// TIA Portal project "CLU" (V13) (continued)
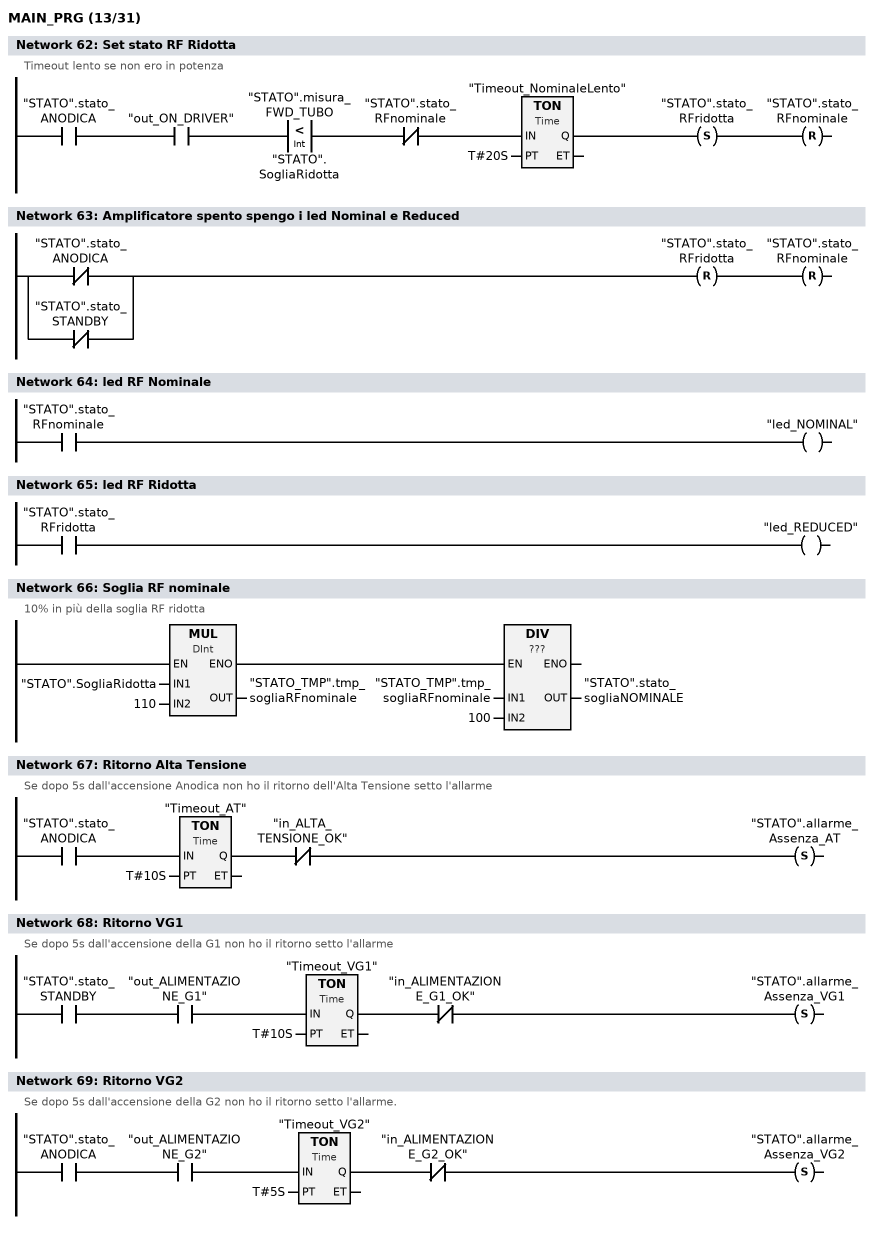
   "Timeout_NominaleLento".TON(IN := "STATO".stato_ANODICA AND "out_ON_DRIVER" AND ("STATO".misura_FWD_TUBO < "STATO".SogliaRidotta) AND NOT "STATO".stato_RFnominale,
                           PT := T#20S);
   IF "Timeout_NominaleLento".Q THEN
       "STATO".stato_RFridotta := TRUE;
       "STATO".stato_RFnominale := FALSE;
   END_IF;
END_REGION

REGION Network 63: Amplificatore spento spengo i led Nominal e Reduced
   RUNG wire#powerrail
      I_Contact( "STATO".stato_ANODICA )
      wire#w1
      R_Coil( "STATO".stato_RFridotta )
      R_Coil( "STATO".stato_RFnominale )
   END_RUNG
   RUNG wire#powerrail
      I_Contact( "STATO".stato_STANDBY )
   END_RUNG wire#w1
   // the same network as SCL:
   IF NOT "STATO".stato_ANODICA OR NOT "STATO".stato_STANDBY THEN
       "STATO".stato_RFridotta := FALSE;
       "STATO".stato_RFnominale := FALSE;
   END_IF;
END_REGION

REGION Network 64: led RF Nominale
   RUNG wire#powerrail
      Contact( "STATO".stato_RFnominale )
      Coil( "led_NOMINAL" )
   END_RUNG
   // the same network as SCL:
   "led_NOMINAL" := "STATO".stato_RFnominale;
END_REGION

REGION Network 65: led RF Ridotta
   RUNG wire#powerrail
      Contact( "STATO".stato_RFridotta )
      Coil( "led_REDUCED" )
   END_RUNG
   // the same network as SCL:
   "led_REDUCED" := "STATO".stato_RFridotta;
END_REGION

REGION Network 66: Soglia RF nominale
   // 10% in più della soglia RF ridotta
   RUNG wire#powerrail
      { S7_Templates := "SrcType := DInt" } Mul(in1 := "STATO".SogliaRidotta, in2 := 110, out => "STATO_TMP".tmp_sogliaRFnominale)
      { S7_Templates := "SrcType := ???" } Div(in1 := "STATO_TMP".tmp_sogliaRFnominale, in2 := 100, out => "STATO".stato_sogliaNOMINALE)
   END_RUNG
   // the same network as SCL:
   "STATO_TMP".tmp_sogliaRFnominale := "STATO".SogliaRidotta * 110;
   "STATO".stato_sogliaNOMINALE := "STATO_TMP".tmp_sogliaRFnominale / 100;
END_REGION

REGION Network 67: Ritorno Alta Tensione
   // Se dopo 5s dall'accensione Anodica non ho il ritorno dell'Alta Tensione setto l'allarme
   "Timeout_AT".TON(IN := "STATO".stato_ANODICA, PT := T#10S);
   IF "Timeout_AT".Q AND NOT "in_ALTA_TENSIONE_OK" THEN "STATO".allarme_Assenza_AT := TRUE; END_IF;
END_REGION

REGION Network 68: Ritorno VG1
   // Se dopo 5s dall'accensione della G1 non ho il ritorno setto l'allarme
   "Timeout_VG1".TON(IN := "STATO".stato_STANDBY AND "out_ALIMENTAZIONE_G1", PT := T#10S);
   IF "Timeout_VG1".Q AND NOT "in_ALIMENTAZIONE_G1_OK" THEN "STATO".allarme_Assenza_VG1 := TRUE; END_IF;
END_REGION

REGION Network 69: Ritorno VG2
   // Se dopo 5s dall'accensione della G2 non ho il ritorno setto l'allarme.
   "Timeout_VG2".TON(IN := "STATO".stato_ANODICA AND "out_ALIMENTAZIONE_G2", PT := T#5S);
   IF "Timeout_VG2".Q AND NOT "in_ALIMENTAZIONE_G2_OK" THEN "STATO".allarme_Assenza_VG2 := TRUE; END_IF;
END_REGION

REGION Network 70: Allarme mancanza VG1
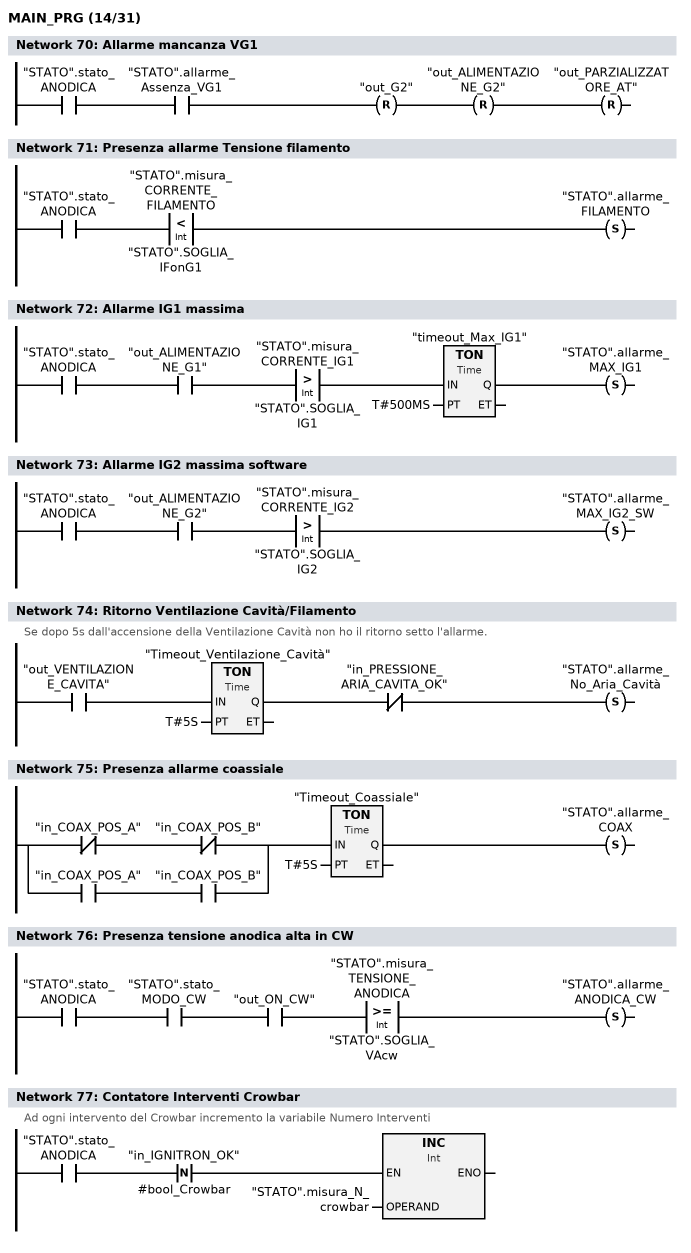
   RUNG wire#powerrail
      Contact( "STATO".stato_ANODICA )
      Contact( "STATO".allarme_Assenza_VG1 )
      R_Coil( "out_G2" )
      R_Coil( "out_ALIMENTAZIONE_G2" )
      R_Coil( "out_PARZIALIZZATORE_AT" )
   END_RUNG
   // the same network as SCL:
   IF "STATO".stato_ANODICA AND "STATO".allarme_Assenza_VG1 THEN
       "out_G2" := FALSE;
       "out_ALIMENTAZIONE_G2" := FALSE;
       "out_PARZIALIZZATORE_AT" := FALSE;
   END_IF;
END_REGION

REGION Network 71: Presenza allarme Tensione filamento
   RUNG wire#powerrail
      Contact( "STATO".stato_ANODICA )
      { S7_Templates := "SrcType := Int" } LT_Contact(in1 := "STATO".misura_CORRENTE_FILAMENTO, in2 := "STATO".SOGLIA_IFonG1)
      S_Coil( "STATO".allarme_FILAMENTO )
   END_RUNG
   // the same network as SCL:
   IF "STATO".stato_ANODICA AND ("STATO".misura_CORRENTE_FILAMENTO < "STATO".SOGLIA_IFonG1) THEN
       "STATO".allarme_FILAMENTO := TRUE;
   END_IF;
END_REGION

REGION Network 72: Allarme IG1 massima
   "timeout_Max_IG1".TON(IN := "STATO".stato_ANODICA AND "out_ALIMENTAZIONE_G1" AND ("STATO".misura_CORRENTE_IG1 > "STATO".SOGLIA_IG1),
                         PT := T#500MS);
   IF "timeout_Max_IG1".Q THEN "STATO".allarme_MAX_IG1 := TRUE; END_IF;
END_REGION

REGION Network 73: Allarme IG2 massima software
   RUNG wire#powerrail
      Contact( "STATO".stato_ANODICA )
      Contact( "out_ALIMENTAZIONE_G2" )
      { S7_Templates := "SrcType := Int" } GT_Contact(in1 := "STATO".misura_CORRENTE_IG2, in2 := "STATO".SOGLIA_IG2)
      S_Coil( "STATO".allarme_MAX_IG2_SW )
   END_RUNG
   // the same network as SCL:
   IF "STATO".stato_ANODICA AND "out_ALIMENTAZIONE_G2" AND ("STATO".misura_CORRENTE_IG2 > "STATO".SOGLIA_IG2) THEN
       "STATO".allarme_MAX_IG2_SW := TRUE;
   END_IF;
END_REGION

REGION Network 74: Ritorno Ventilazione Cavità/Filamento
   // Se dopo 5s dall'accensione della Ventilazione Cavità non ho il ritorno setto l'allarme.
   "Timeout_Ventilazione_Cavità".TON(IN := "out_VENTILAZIONE_CAVITA", PT := T#5S);
   IF "Timeout_Ventilazione_Cavità".Q AND NOT "in_PRESSIONE_ARIA_CAVITA_OK" THEN
       "STATO".allarme_No_Aria_Cavità := TRUE;
   END_IF;
END_REGION

REGION Network 75: Presenza allarme coassiale
   "Timeout_Coassiale".TON(IN := (NOT "in_COAX_POS_A" AND NOT "in_COAX_POS_B") OR ("in_COAX_POS_A" AND "in_COAX_POS_B"),
                           PT := T#5S);
   IF "Timeout_Coassiale".Q THEN "STATO".allarme_COAX := TRUE; END_IF;
END_REGION

REGION Network 76: Presenza tensione anodica alta in CW
   RUNG wire#powerrail
      Contact( "STATO".stato_ANODICA )
      Contact( "STATO".stato_MODO_CW )
      Contact( "out_ON_CW" )
      { S7_Templates := "SrcType := Int" } GE_Contact(in1 := "STATO".misura_TENSIONE_ANODICA, in2 := "STATO".SOGLIA_VAcw)
      S_Coil( "STATO".allarme_ANODICA_CW )
   END_RUNG
   // the same network as SCL:
   IF "STATO".stato_ANODICA AND "STATO".stato_MODO_CW AND "out_ON_CW" AND ("STATO".misura_TENSIONE_ANODICA >= "STATO".SOGLIA_VAcw) THEN
       "STATO".allarme_ANODICA_CW := TRUE;
   END_IF;
END_REGION

REGION Network 77: Contatore Interventi Crowbar
   // Ad ogni intervento del Crowbar incremento la variabile Numero Interventi
   RUNG wire#powerrail
      Contact( "STATO".stato_ANODICA )
      N_Contact(operand := "in_IGNITRON_OK", bit := #bool_Crowbar)
      { S7_Templates := "DestType := Int" } Inc( "STATO".misura_N_crowbar )
   END_RUNG
   // the same network as SCL:
   #_w1 := "STATO".stato_ANODICA AND NOT "in_IGNITRON_OK" AND #bool_Crowbar;   // falling edge of "in_IGNITRON_OK"
   #bool_Crowbar := "in_IGNITRON_OK";
   IF #_w1 THEN "STATO".misura_N_crowbar := "STATO".misura_N_crowbar + 1; END_IF;
END_REGION

REGION Network 78: Soglia ROS 400kW
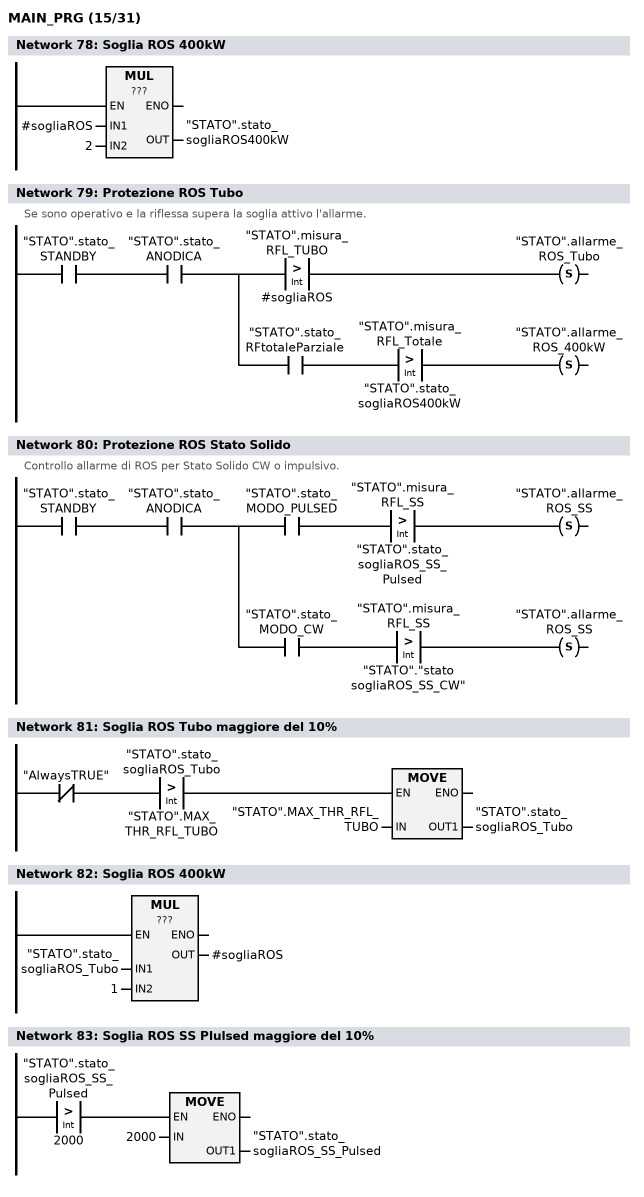
   RUNG wire#powerrail
      { S7_Templates := "SrcType := ???" } Mul(in1 := #sogliaROS, in2 := 2, out => "STATO".stato_sogliaROS400kW)
   END_RUNG
   // the same network as SCL:
   "STATO".stato_sogliaROS400kW := #sogliaROS * 2;
END_REGION

REGION Network 79: Protezione ROS Tubo
   // Se sono operativo e la riflessa supera la soglia attivo l'allarme.
   RUNG wire#powerrail
      Contact( "STATO".stato_STANDBY )
      Contact( "STATO".stato_ANODICA )
      wire#w1
      { S7_Templates := "SrcType := Int" } GT_Contact(in1 := "STATO".misura_RFL_TUBO, in2 := #sogliaROS)
      S_Coil( "STATO".allarme_ROS_Tubo )
   END_RUNG
   RUNG wire#w1
      Contact( "STATO".stato_RFtotaleParziale )
      { S7_Templates := "SrcType := Int" } GT_Contact(in1 := "STATO".misura_RFL_Totale, in2 := "STATO".stato_sogliaROS400kW)
      S_Coil( "STATO".allarme_ROS_400kW )
   END_RUNG
   // the same network as SCL:
   #_w1 := "STATO".stato_STANDBY AND "STATO".stato_ANODICA;
   IF #_w1 AND ("STATO".misura_RFL_TUBO > #sogliaROS) THEN "STATO".allarme_ROS_Tubo := TRUE; END_IF;
   IF #_w1 AND "STATO".stato_RFtotaleParziale AND ("STATO".misura_RFL_Totale > "STATO".stato_sogliaROS400kW) THEN
       "STATO".allarme_ROS_400kW := TRUE;
   END_IF;
END_REGION

REGION Network 80: Protezione ROS Stato Solido
   // Controllo allarme di ROS per Stato Solido CW o impulsivo.
   RUNG wire#powerrail
      Contact( "STATO".stato_STANDBY )
      Contact( "STATO".stato_ANODICA )
      wire#w1
      Contact( "STATO".stato_MODO_PULSED )
      { S7_Templates := "SrcType := Int" } GT_Contact(in1 := "STATO".misura_RFL_SS, in2 := "STATO".stato_sogliaROS_SS_Pulsed)
      S_Coil( "STATO".allarme_ROS_SS )
   END_RUNG
   RUNG wire#w1
      Contact( "STATO".stato_MODO_CW )
      { S7_Templates := "SrcType := Int" } GT_Contact(in1 := "STATO".misura_RFL_SS, in2 := "STATO"."stato sogliaROS_SS_CW")
      S_Coil( "STATO".allarme_ROS_SS )
   END_RUNG
   // the same network as SCL:
   #_w1 := "STATO".stato_STANDBY AND "STATO".stato_ANODICA;
   IF #_w1 AND "STATO".stato_MODO_PULSED AND ("STATO".misura_RFL_SS > "STATO".stato_sogliaROS_SS_Pulsed) THEN
       "STATO".allarme_ROS_SS := TRUE;
   END_IF;
   IF #_w1 AND "STATO".stato_MODO_CW AND ("STATO".misura_RFL_SS > "STATO"."stato sogliaROS_SS_CW") THEN
       "STATO".allarme_ROS_SS := TRUE;
   END_IF;
END_REGION

REGION Network 81: Soglia ROS Tubo maggiore del 10%
   RUNG wire#powerrail
      I_Contact( "AlwaysTRUE" )
      { S7_Templates := "SrcType := Int" } GT_Contact(in1 := "STATO".stato_sogliaROS_Tubo, in2 := "STATO".MAX_THR_RFL_TUBO)
      Move(in := "STATO".MAX_THR_RFL_TUBO, out1 => "STATO".stato_sogliaROS_Tubo)
   END_RUNG
   // the same network as SCL:
   IF NOT "AlwaysTRUE" AND ("STATO".stato_sogliaROS_Tubo > "STATO".MAX_THR_RFL_TUBO) THEN
       "STATO".stato_sogliaROS_Tubo := "STATO".MAX_THR_RFL_TUBO;
   END_IF;
END_REGION

REGION Network 82: Soglia ROS 400kW
   RUNG wire#powerrail
      { S7_Templates := "SrcType := ???" } Mul(in1 := "STATO".stato_sogliaROS_Tubo, in2 := 1, out => #sogliaROS)
   END_RUNG
   // the same network as SCL:
   #sogliaROS := "STATO".stato_sogliaROS_Tubo * 1;
END_REGION

REGION Network 83: Soglia ROS SS Plulsed maggiore del 10%
   RUNG wire#powerrail
      { S7_Templates := "SrcType := Int" } GT_Contact(in1 := "STATO".stato_sogliaROS_SS_Pulsed, in2 := 2000)
      Move(in := 2000, out1 => "STATO".stato_sogliaROS_SS_Pulsed)
   END_RUNG
   // the same network as SCL:
   IF "STATO".stato_sogliaROS_SS_Pulsed > 2000 THEN "STATO".stato_sogliaROS_SS_Pulsed := 2000; END_IF;
END_REGION

REGION Network 84: Soglia ROS SS CW maggiore del 10%
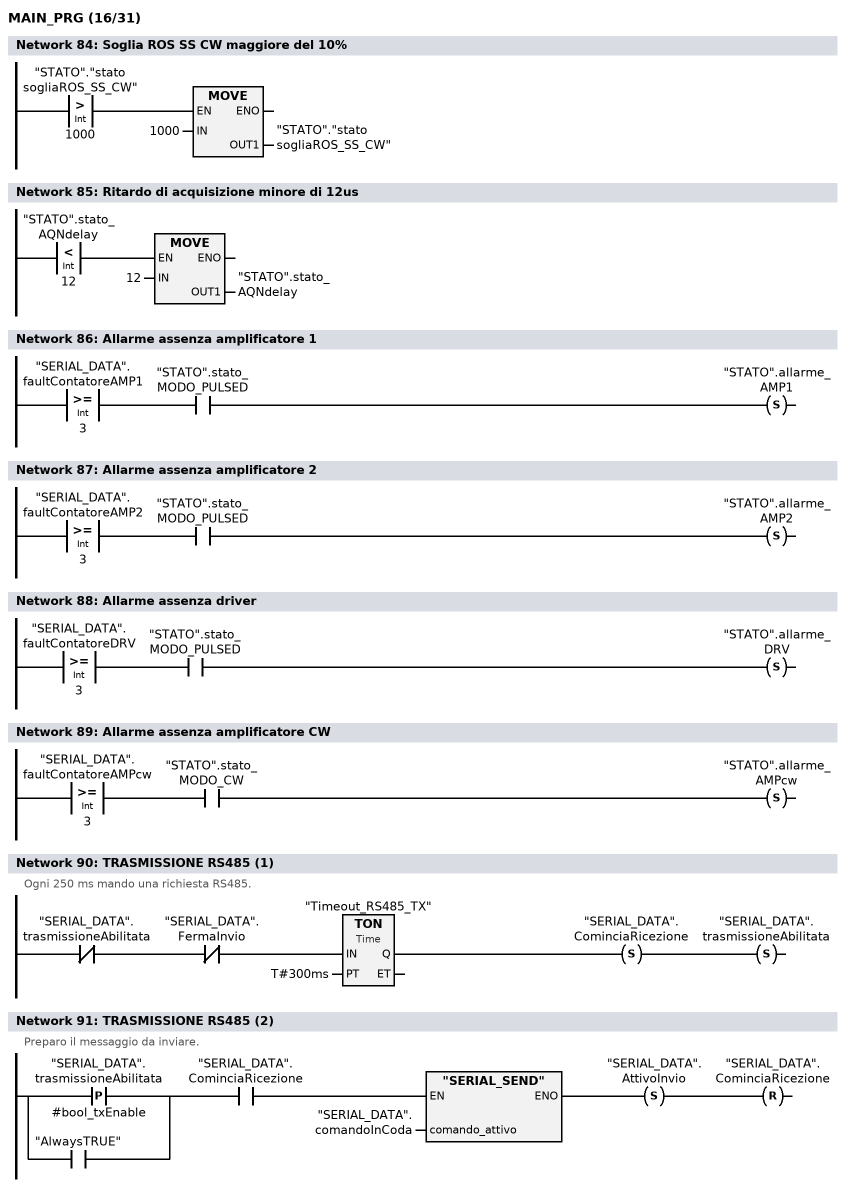
   RUNG wire#powerrail
      { S7_Templates := "SrcType := Int" } GT_Contact(in1 := "STATO"."stato sogliaROS_SS_CW", in2 := 1000)
      Move(in := 1000, out1 => "STATO"."stato sogliaROS_SS_CW")
   END_RUNG
   // the same network as SCL:
   IF "STATO"."stato sogliaROS_SS_CW" > 1000 THEN "STATO"."stato sogliaROS_SS_CW" := 1000; END_IF;
END_REGION

REGION Network 85: Ritardo di acquisizione minore di 12us
   RUNG wire#powerrail
      { S7_Templates := "SrcType := Int" } LT_Contact(in1 := "STATO".stato_AQNdelay, in2 := 12)
      Move(in := 12, out1 => "STATO".stato_AQNdelay)
   END_RUNG
   // the same network as SCL:
   IF "STATO".stato_AQNdelay < 12 THEN "STATO".stato_AQNdelay := 12; END_IF;
END_REGION

REGION Network 86: Allarme assenza amplificatore 1
   RUNG wire#powerrail
      { S7_Templates := "SrcType := Int" } GE_Contact(in1 := "SERIAL_DATA".faultContatoreAMP1, in2 := 3)
      Contact( "STATO".stato_MODO_PULSED )
      S_Coil( "STATO".allarme_AMP1 )
   END_RUNG
   // the same network as SCL:
   IF ("SERIAL_DATA".faultContatoreAMP1 >= 3) AND "STATO".stato_MODO_PULSED THEN
       "STATO".allarme_AMP1 := TRUE;
   END_IF;
END_REGION

REGION Network 87: Allarme assenza amplificatore 2
   RUNG wire#powerrail
      { S7_Templates := "SrcType := Int" } GE_Contact(in1 := "SERIAL_DATA".faultContatoreAMP2, in2 := 3)
      Contact( "STATO".stato_MODO_PULSED )
      S_Coil( "STATO".allarme_AMP2 )
   END_RUNG
   // the same network as SCL:
   IF ("SERIAL_DATA".faultContatoreAMP2 >= 3) AND "STATO".stato_MODO_PULSED THEN
       "STATO".allarme_AMP2 := TRUE;
   END_IF;
END_REGION

REGION Network 88: Allarme assenza driver
   RUNG wire#powerrail
      { S7_Templates := "SrcType := Int" } GE_Contact(in1 := "SERIAL_DATA".faultContatoreDRV, in2 := 3)
      Contact( "STATO".stato_MODO_PULSED )
      S_Coil( "STATO".allarme_DRV )
   END_RUNG
   // the same network as SCL:
   IF ("SERIAL_DATA".faultContatoreDRV >= 3) AND "STATO".stato_MODO_PULSED THEN
       "STATO".allarme_DRV := TRUE;
   END_IF;
END_REGION

REGION Network 89: Allarme assenza amplificatore CW
   RUNG wire#powerrail
      { S7_Templates := "SrcType := Int" } GE_Contact(in1 := "SERIAL_DATA".faultContatoreAMPcw, in2 := 3)
      Contact( "STATO".stato_MODO_CW )
      S_Coil( "STATO".allarme_AMPcw )
   END_RUNG
   // the same network as SCL:
   IF ("SERIAL_DATA".faultContatoreAMPcw >= 3) AND "STATO".stato_MODO_CW THEN
       "STATO".allarme_AMPcw := TRUE;
   END_IF;
END_REGION

REGION Network 90: TRASMISSIONE RS485 (1)
   // Ogni 250 ms mando una richiesta RS485.
   "Timeout_RS485_TX".TON(IN := NOT "SERIAL_DATA".trasmissioneAbilitata AND NOT "SERIAL_DATA".FermaInvio,
                          PT := T#300ms);
   IF "Timeout_RS485_TX".Q THEN
       "SERIAL_DATA".CominciaRicezione := TRUE;
       "SERIAL_DATA".trasmissioneAbilitata := TRUE;
   END_IF;
END_REGION

REGION Network 91: TRASMISSIONE RS485 (2)
   // Preparo il messaggio da inviare.
   RUNG wire#powerrail
      P_Contact(operand := "SERIAL_DATA".trasmissioneAbilitata, bit := #bool_txEnable)
      wire#w1
      Contact( "SERIAL_DATA".CominciaRicezione )
      "SERIAL_SEND"(comando_attivo := "SERIAL_DATA".comandoInCoda)
      S_Coil( "SERIAL_DATA".AttivoInvio )
      R_Coil( "SERIAL_DATA".CominciaRicezione )
   END_RUNG
   RUNG wire#powerrail
      Contact( "AlwaysTRUE" )
   END_RUNG wire#w1
   // the same network as SCL:
   #_w1 := "SERIAL_DATA".trasmissioneAbilitata AND NOT #bool_txEnable;   // rising edge of "SERIAL_DATA".trasmissioneAbilitata
   #bool_txEnable := "SERIAL_DATA".trasmissioneAbilitata;
   "SERIAL_SEND"(EN := (#_w1 OR "AlwaysTRUE") AND "SERIAL_DATA".CominciaRicezione,
                 comando_attivo := "SERIAL_DATA".comandoInCoda,
                 ENO => #_w2);
   IF #_w2 THEN
       "SERIAL_DATA".AttivoInvio := TRUE;
       "SERIAL_DATA".CominciaRicezione := FALSE;
   END_IF;
END_REGION

REGION Network 92: TRASMISSIONE RS485 (3): 76h
   // Processo la richiesta di stato ID==0
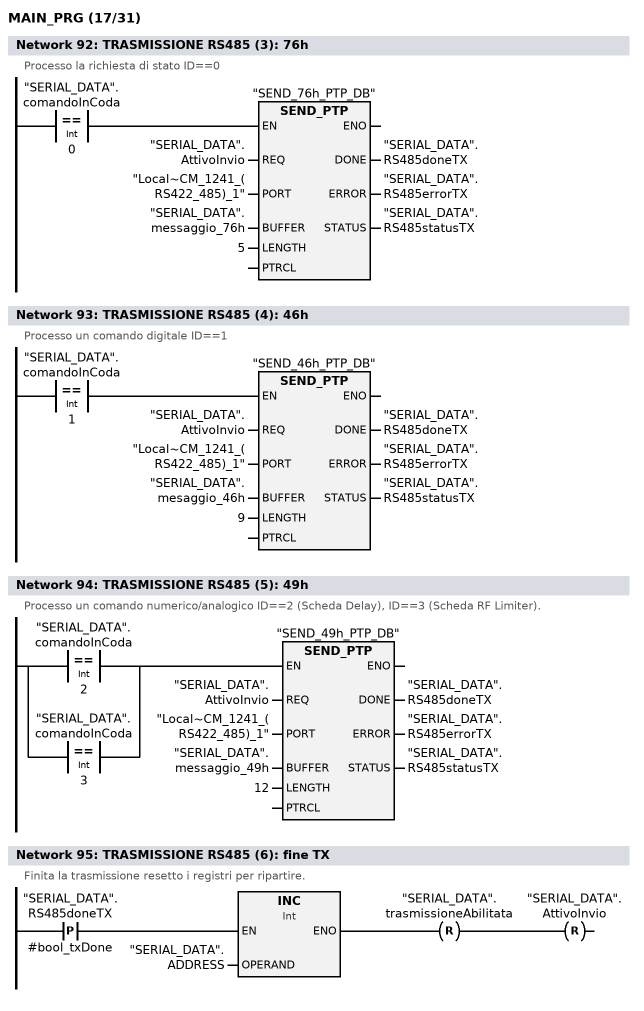
   IF "SERIAL_DATA".comandoInCoda = 0 THEN
       "SEND_76h_PTP_DB"(REQ := "SERIAL_DATA".AttivoInvio,   // SEND_PTP
                         PORT := "Local~CM_1241_(RS422_485)_1",
                         BUFFER := "SERIAL_DATA".messaggio_76h,
                         LENGTH := 5,
                         DONE => "SERIAL_DATA".RS485doneTX,
                         ERROR => "SERIAL_DATA".RS485errorTX,
                         STATUS => "SERIAL_DATA".RS485statusTX);
   END_IF;
END_REGION

REGION Network 93: TRASMISSIONE RS485 (4): 46h
   // Processo un comando digitale ID==1
   IF "SERIAL_DATA".comandoInCoda = 1 THEN
       "SEND_46h_PTP_DB"(REQ := "SERIAL_DATA".AttivoInvio,   // SEND_PTP
                         PORT := "Local~CM_1241_(RS422_485)_1",
                         BUFFER := "SERIAL_DATA".mesaggio_46h,
                         LENGTH := 9,
                         DONE => "SERIAL_DATA".RS485doneTX,
                         ERROR => "SERIAL_DATA".RS485errorTX,
                         STATUS => "SERIAL_DATA".RS485statusTX);
   END_IF;
END_REGION

REGION Network 94: TRASMISSIONE RS485 (5): 49h
   // Processo un comando numerico/analogico ID==2 (Scheda Delay), ID==3 (Scheda RF Limiter).
   IF ("SERIAL_DATA".comandoInCoda = 2) OR ("SERIAL_DATA".comandoInCoda = 3) THEN
       "SEND_49h_PTP_DB"(REQ := "SERIAL_DATA".AttivoInvio,   // SEND_PTP
                         PORT := "Local~CM_1241_(RS422_485)_1",
                         BUFFER := "SERIAL_DATA".messaggio_49h,
                         LENGTH := 12,
                         DONE => "SERIAL_DATA".RS485doneTX,
                         ERROR => "SERIAL_DATA".RS485errorTX,
                         STATUS => "SERIAL_DATA".RS485statusTX);
   END_IF;
END_REGION

REGION Network 95: TRASMISSIONE RS485 (6): fine TX
   // Finita la trasmissione resetto i registri per ripartire.
   RUNG wire#powerrail
      P_Contact(operand := "SERIAL_DATA".RS485doneTX, bit := #bool_txDone)
      { S7_Templates := "DestType := Int" } Inc( "SERIAL_DATA".ADDRESS )
      R_Coil( "SERIAL_DATA".trasmissioneAbilitata )
      R_Coil( "SERIAL_DATA".AttivoInvio )
   END_RUNG
   // the same network as SCL:
   #_w1 := "SERIAL_DATA".RS485doneTX AND NOT #bool_txDone;   // rising edge of "SERIAL_DATA".RS485doneTX
   #bool_txDone := "SERIAL_DATA".RS485doneTX;
   IF #_w1 THEN
       "SERIAL_DATA".ADDRESS := "SERIAL_DATA".ADDRESS + 1;
       "SERIAL_DATA".trasmissioneAbilitata := FALSE;
       "SERIAL_DATA".AttivoInvio := FALSE;
   END_IF;
END_REGION

REGION Network 96: RICEZIONE RS485 (1): ricezione
   // La ricezione seriale è sempre attiva.
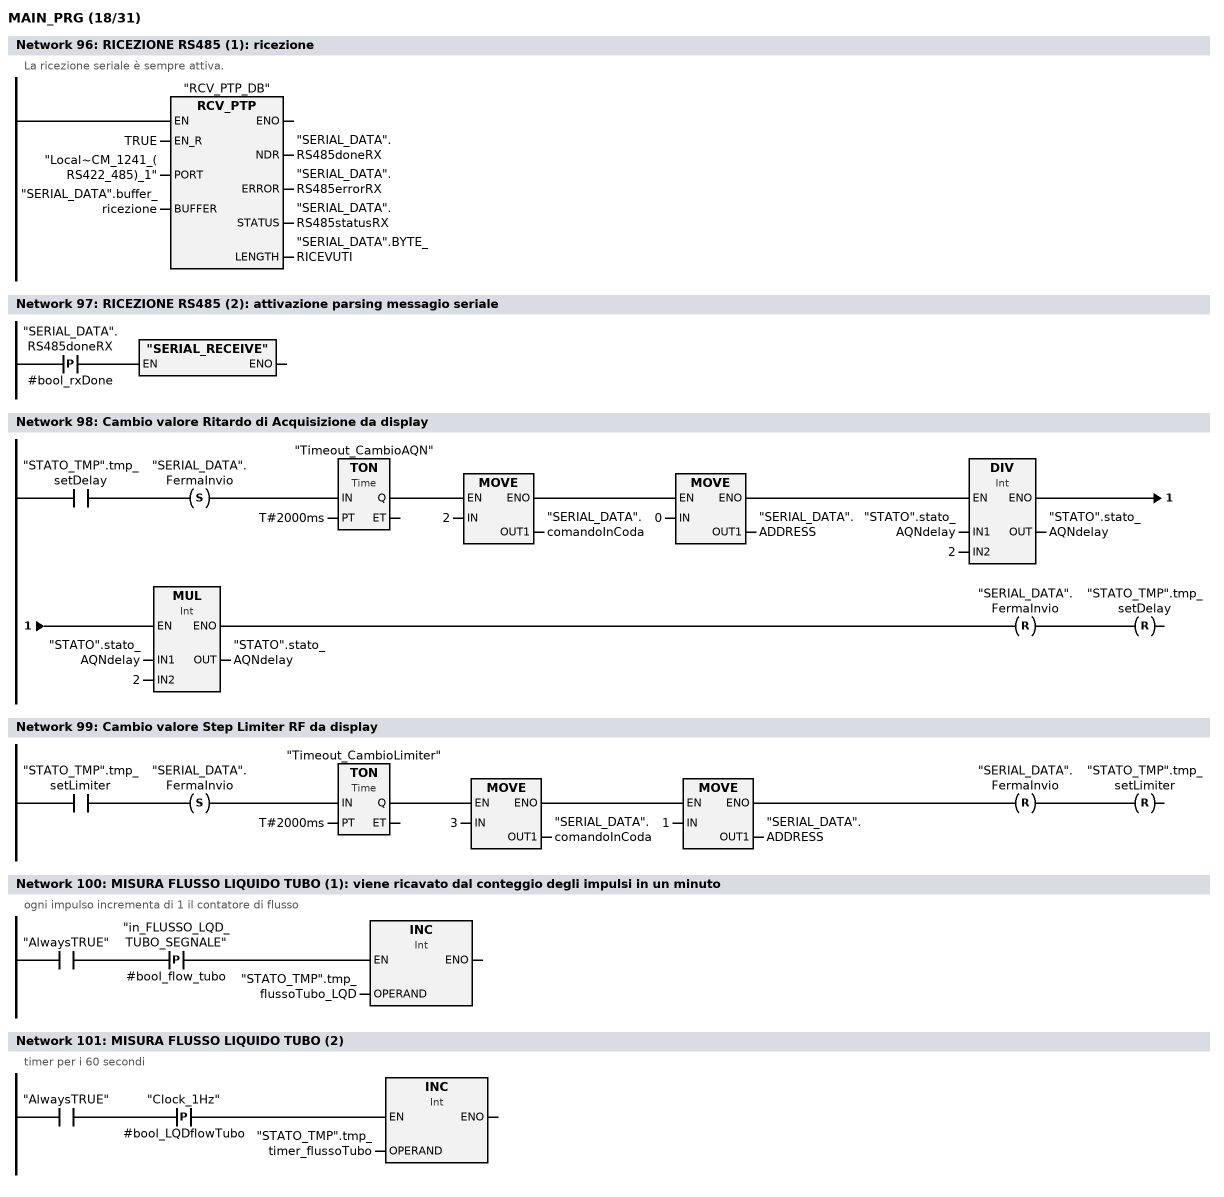
   "RCV_PTP_DB"(EN_R := TRUE,   // RCV_PTP
                PORT := "Local~CM_1241_(RS422_485)_1",
                BUFFER := "SERIAL_DATA".buffer_ricezione,
                NDR => "SERIAL_DATA".RS485doneRX,
                ERROR => "SERIAL_DATA".RS485errorRX,
                STATUS => "SERIAL_DATA".RS485statusRX,
                LENGTH => "SERIAL_DATA".BYTE_RICEVUTI);
END_REGION

REGION Network 97: RICEZIONE RS485 (2): attivazione parsing messagio seriale
   RUNG wire#powerrail
      P_Contact(operand := "SERIAL_DATA".RS485doneRX, bit := #bool_rxDone)
      "SERIAL_RECEIVE"()
   END_RUNG
   // the same network as SCL:
   #_w1 := "SERIAL_DATA".RS485doneRX AND NOT #bool_rxDone;   // rising edge of "SERIAL_DATA".RS485doneRX
   #bool_rxDone := "SERIAL_DATA".RS485doneRX;
   IF #_w1 THEN "SERIAL_RECEIVE"(); END_IF;
END_REGION

REGION Network 98: Cambio valore Ritardo di Acquisizione da display
   IF "STATO_TMP".tmp_setDelay THEN "SERIAL_DATA".FermaInvio := TRUE; END_IF;
   "Timeout_CambioAQN".TON(IN := "STATO_TMP".tmp_setDelay, PT := T#2000ms);
   IF "Timeout_CambioAQN".Q THEN
       "SERIAL_DATA".comandoInCoda := 2;
       "SERIAL_DATA".ADDRESS := 0;
       "STATO".stato_AQNdelay := "STATO".stato_AQNdelay / 2;
       "STATO".stato_AQNdelay := "STATO".stato_AQNdelay * 2;
       "SERIAL_DATA".FermaInvio := FALSE;
       "STATO_TMP".tmp_setDelay := FALSE;
   END_IF;
END_REGION

REGION Network 99: Cambio valore Step Limiter RF da display
   IF "STATO_TMP".tmp_setLimiter THEN "SERIAL_DATA".FermaInvio := TRUE; END_IF;
   "Timeout_CambioLimiter".TON(IN := "STATO_TMP".tmp_setLimiter, PT := T#2000ms);
   IF "Timeout_CambioLimiter".Q THEN
       "SERIAL_DATA".comandoInCoda := 3;
       "SERIAL_DATA".ADDRESS := 1;
       "SERIAL_DATA".FermaInvio := FALSE;
       "STATO_TMP".tmp_setLimiter := FALSE;
   END_IF;
END_REGION

REGION Network 100: MISURA FLUSSO LIQUIDO TUBO (1): viene ricavato dal conteggio degli impulsi in un minuto
   // ogni impulso incrementa di 1 il contatore di flusso
   RUNG wire#powerrail
      Contact( "AlwaysTRUE" )
      P_Contact(operand := "in_FLUSSO_LQD_TUBO_SEGNALE", bit := #bool_flow_tubo)
      { S7_Templates := "DestType := Int" } Inc( "STATO_TMP".tmp_flussoTubo_LQD )
   END_RUNG
   // the same network as SCL:
   #_w1 := "AlwaysTRUE" AND "in_FLUSSO_LQD_TUBO_SEGNALE" AND NOT #bool_flow_tubo;   // rising edge of "in_FLUSSO_LQD_TUBO_SEGNALE"
   #bool_flow_tubo := "in_FLUSSO_LQD_TUBO_SEGNALE";
   IF #_w1 THEN "STATO_TMP".tmp_flussoTubo_LQD := "STATO_TMP".tmp_flussoTubo_LQD + 1; END_IF;
END_REGION

REGION Network 101: MISURA FLUSSO LIQUIDO TUBO (2)
   // timer per i 60 secondi
   RUNG wire#powerrail
      Contact( "AlwaysTRUE" )
      P_Contact(operand := "Clock_1Hz", bit := #bool_LQDflowTubo)
      { S7_Templates := "DestType := Int" } Inc( "STATO_TMP".tmp_timer_flussoTubo )
   END_RUNG
   // the same network as SCL:
   #_w1 := "AlwaysTRUE" AND "Clock_1Hz" AND NOT #bool_LQDflowTubo;   // rising edge of "Clock_1Hz"
   #bool_LQDflowTubo := "Clock_1Hz";
   IF #_w1 THEN "STATO_TMP".tmp_timer_flussoTubo := "STATO_TMP".tmp_timer_flussoTubo + 1; END_IF;
END_REGION

REGION Network 102: MISURA FLUSSO LIQUIDO TUBO (3)
   // dopo 60 secondi calcolo scalo la misura
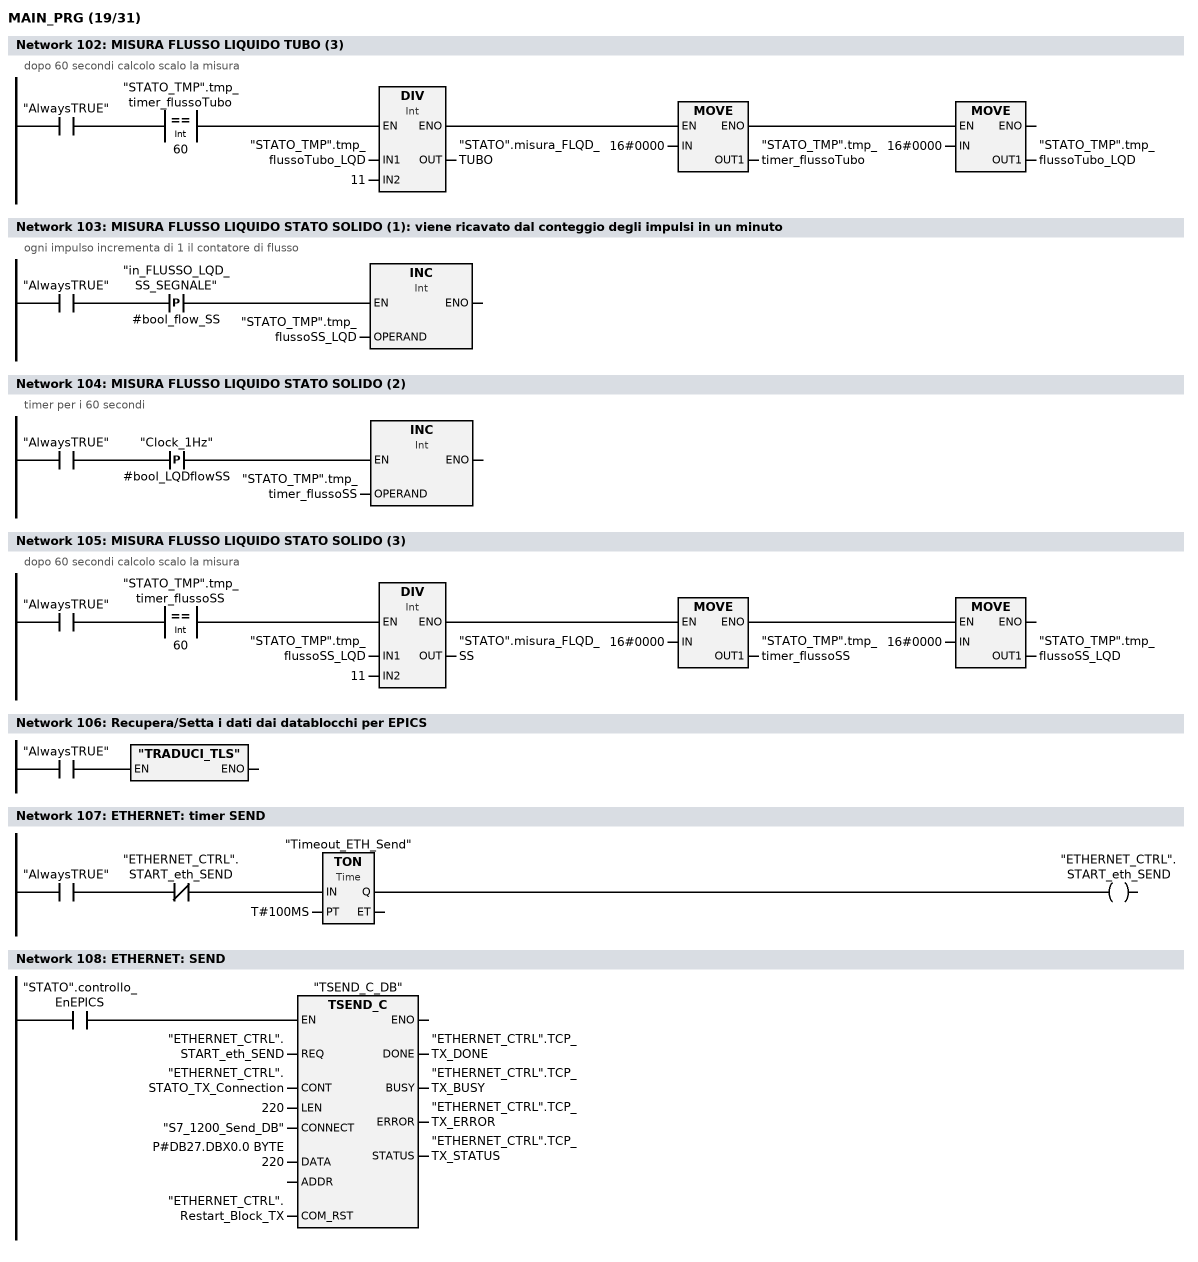
   RUNG wire#powerrail
      Contact( "AlwaysTRUE" )
      { S7_Templates := "SrcType := Int" } EQ_Contact(in1 := "STATO_TMP".tmp_timer_flussoTubo, in2 := 60)
      { S7_Templates := "SrcType := Int" } Div(in1 := "STATO_TMP".tmp_flussoTubo_LQD, in2 := 11, out => "STATO".misura_FLQD_TUBO)
      { S7_GenerateENO := "TRUE" } Move(in := 16#0000, out1 => "STATO_TMP".tmp_timer_flussoTubo)
      { S7_GenerateENO := "TRUE" } Move(in := 16#0000, out1 => "STATO_TMP".tmp_flussoTubo_LQD)
   END_RUNG
   // the same network as SCL:
   // ENO of a box is taken as its EN; it also drops when the box reports an error
   IF "AlwaysTRUE" AND ("STATO_TMP".tmp_timer_flussoTubo = 60) THEN
       "STATO".misura_FLQD_TUBO := "STATO_TMP".tmp_flussoTubo_LQD / 11;
   END_IF;
   #_w1 := "AlwaysTRUE" AND ("STATO_TMP".tmp_timer_flussoTubo = 60);
   IF #_w1 THEN
       "STATO_TMP".tmp_timer_flussoTubo := 16#0000;
       "STATO_TMP".tmp_flussoTubo_LQD := 16#0000;
   END_IF;
END_REGION

REGION Network 103: MISURA FLUSSO LIQUIDO STATO SOLIDO (1): viene ricavato dal conteggio degli impulsi in un minuto
   // ogni impulso incrementa di 1 il contatore di flusso
   RUNG wire#powerrail
      Contact( "AlwaysTRUE" )
      P_Contact(operand := "in_FLUSSO_LQD_SS_SEGNALE", bit := #bool_flow_SS)
      { S7_Templates := "DestType := Int" } Inc( "STATO_TMP".tmp_flussoSS_LQD )
   END_RUNG
   // the same network as SCL:
   #_w1 := "AlwaysTRUE" AND "in_FLUSSO_LQD_SS_SEGNALE" AND NOT #bool_flow_SS;   // rising edge of "in_FLUSSO_LQD_SS_SEGNALE"
   #bool_flow_SS := "in_FLUSSO_LQD_SS_SEGNALE";
   IF #_w1 THEN "STATO_TMP".tmp_flussoSS_LQD := "STATO_TMP".tmp_flussoSS_LQD + 1; END_IF;
END_REGION

REGION Network 104: MISURA FLUSSO LIQUIDO STATO SOLIDO (2)
   // timer per i 60 secondi
   RUNG wire#powerrail
      Contact( "AlwaysTRUE" )
      P_Contact(operand := "Clock_1Hz", bit := #bool_LQDflowSS)
      { S7_Templates := "DestType := Int" } Inc( "STATO_TMP".tmp_timer_flussoSS )
   END_RUNG
   // the same network as SCL:
   #_w1 := "AlwaysTRUE" AND "Clock_1Hz" AND NOT #bool_LQDflowSS;   // rising edge of "Clock_1Hz"
   #bool_LQDflowSS := "Clock_1Hz";
   IF #_w1 THEN "STATO_TMP".tmp_timer_flussoSS := "STATO_TMP".tmp_timer_flussoSS + 1; END_IF;
END_REGION

REGION Network 105: MISURA FLUSSO LIQUIDO STATO SOLIDO (3)
   // dopo 60 secondi calcolo scalo la misura
   RUNG wire#powerrail
      Contact( "AlwaysTRUE" )
      { S7_Templates := "SrcType := Int" } EQ_Contact(in1 := "STATO_TMP".tmp_timer_flussoSS, in2 := 60)
      { S7_Templates := "SrcType := Int" } Div(in1 := "STATO_TMP".tmp_flussoSS_LQD, in2 := 11, out => "STATO".misura_FLQD_SS)
      { S7_GenerateENO := "TRUE" } Move(in := 16#0000, out1 => "STATO_TMP".tmp_timer_flussoSS)
      { S7_GenerateENO := "TRUE" } Move(in := 16#0000, out1 => "STATO_TMP".tmp_flussoSS_LQD)
   END_RUNG
   // the same network as SCL:
   // ENO of a box is taken as its EN; it also drops when the box reports an error
   IF "AlwaysTRUE" AND ("STATO_TMP".tmp_timer_flussoSS = 60) THEN
       "STATO".misura_FLQD_SS := "STATO_TMP".tmp_flussoSS_LQD / 11;
   END_IF;
   #_w1 := "AlwaysTRUE" AND ("STATO_TMP".tmp_timer_flussoSS = 60);
   IF #_w1 THEN
       "STATO_TMP".tmp_timer_flussoSS := 16#0000;
       "STATO_TMP".tmp_flussoSS_LQD := 16#0000;
   END_IF;
END_REGION

REGION Network 106: Recupera/Setta i dati dai datablocchi per EPICS
   RUNG wire#powerrail
      Contact( "AlwaysTRUE" )
      "TRADUCI_TLS"()
   END_RUNG
   // the same network as SCL:
   IF "AlwaysTRUE" THEN "TRADUCI_TLS"(); END_IF;
END_REGION

REGION Network 107: ETHERNET: timer SEND
   "Timeout_ETH_Send".TON(IN := "AlwaysTRUE" AND NOT "ETHERNET_CTRL".START_eth_SEND, PT := T#100MS);
   "ETHERNET_CTRL".START_eth_SEND := "Timeout_ETH_Send".Q;
END_REGION

REGION Network 108: ETHERNET: SEND
   IF "STATO".controllo_EnEPICS THEN
       "TSEND_C_DB"(REQ := "ETHERNET_CTRL".START_eth_SEND,   // TSEND_C
                    CONT := "ETHERNET_CTRL".STATO_TX_Connection,
                    LEN := 220,
                    CONNECT := "S7_1200_Send_DB",
                    DATA := P#DB27.DBX0.0 BYTE 220,
                    COM_RST := "ETHERNET_CTRL".Restart_Block_TX,
                    DONE => "ETHERNET_CTRL".TCP_TX_DONE,
                    BUSY => "ETHERNET_CTRL".TCP_TX_BUSY,
                    ERROR => "ETHERNET_CTRL".TCP_TX_ERROR,
                    STATUS => "ETHERNET_CTRL".TCP_TX_STATUS);
   END_IF;
END_REGION

